(* Logix 5000 project; controller PLC_MCC1300_75F1 vendor 1 type 14 code 166 rev 32.11; software revision 32.04; part 76 of 83 *)
(* tags used below, declared in another part *)
   AUX_tCapsConveyor_NULL : UDT_CapsConveyor_ZC;
   CONST_tPlant : UDT_PLANT_CONSTANTS;
   M302SpeedUp_ALM : MAC_SpeedUp_ALM;
   M307ASpeedUp_ALM : MAC_SpeedUp_ALM;
   M30xTrimDeck : MAC_TrimmingDeck[5];
   M30xTrimWheel : MAC_TrimmingWheels[5];
   M312 : MAC_Conveyor_Single;
   TMP_dIndex : DINT;
   TMP_dIndexCapConv : DINT;
   TMP_dIndexConv : DINT;
   TMP_x : BOOL;
   TMP_xDummy : BOOL;
   xAlwaysOFF : BOOL;
   Z300_BufferPlate : UDT_LINE_BUFFER_PLATE;
   Z300_Conveyor : UDT_StandConv[29];
   Z300_Conveyor_HMW : MAC_Conveyor_ZC_HMW[29];
   Z300_LineTracking : UDT_LINE_TRACKING;
   Z301 : MAC_Zone_ML;
   Z301_ALM : MAC_Zone_ML_ALM;
   Z301_HMR : MAC_Zone_ML_HMR;
   Z301_HMW : MAC_Zone_ML_HMW;
(* MainProgram, continued *)

ROUTINE Tracking_Logic   (* structured text *)
   
   // Step advancement conveyor
   FOR TMP_dIndexConv:=0 TO CONST_tPlant.dNumOfConveyors - 1 DO
   	JSR(sbrTrackingConvStep,1,TMP_dIndexConv);
   	//reset conveyor tracking
   	FOR TMP_dIndexCapConv := 0 TO CONST_tPlant.dNumCapsConveyor - 1 DO
   		COP(AUX_tCapsConveyor_NULL,Z300_LineTracking.rgtTrkConv[TMP_dIndexConv].Cap[TMP_dIndexCapConv],1);
   	END_FOR;
   	Z300_LineTracking.rgtTrkConv[TMP_dIndexConv].dIndexCaps := 0;
   	Z300_LineTracking.rgtTrkConv[TMP_dIndexConv].xPlatePassageNext := 0;
   	Z300_LineTracking.rgtTrkConv[TMP_dIndexConv].xPlatePassagePrevious := 0;
   	Z300_LineTracking.rgtTrkConv[TMP_dIndexConv].xGlassPresence := 0;
   	Z300_LineTracking.rgtTrkConv[TMP_dIndexConv].xPlateConvPreviousNext := 0;
   	Z300_LineTracking.rgtTrkConv[TMP_dIndexConv].dTailPosition_cmm := 0;
   	Z300_LineTracking.rgtTrkConv[TMP_dIndexConv].dHeadPosition_cmm := 0;
   END_FOR;
   
   // Reset flag for tracking
   FOR TMP_dIndex:=0 TO CONST_tPlant.dMaxNumPlates - 1 DO
   	IF Z300_BufferPlate.rgtPlate[TMP_dIndex].tData.dLength_cmm <= 0 THEN
   		Z300_BufferPlate.rgtPlate[TMP_dIndex].tTracking.xHoldAdvancement := 0;
   		Z300_BufferPlate.rgtPlate[TMP_dIndex].tTracking.xNotConsConvTrk := 0;
   		Z300_BufferPlate.rgtPlate[TMP_dIndex].tTracking.xNotShownInScada := 0;
   	END_IF;
   END_FOR;
   
   // Tracking index not in convoy
   FOR TMP_dIndex:=0 TO CONST_tPlant.dMaxNumPlates - 1 DO
   	JSR(sbrTrackingIndexNotInConvoy,1,Z300_BufferPlate.rgtPlate[TMP_dIndex].tTracking);
   END_FOR;
   
   // Tracking shift
   JSR(sbrTrackingShift);
   
   // Plate presence convoy
   JSR(sbrTrackingConvPresence);
   
END_ROUTINE

ROUTINE Z301_Faults   (* ladder *)
   0: NOP();
   1: XIC(Z301.ST_xAlarmOff)MOV(0,Z301_ALM.rgxEmergency[0])MOV(0,Z301_ALM.rgxStoppingFault[0])MOV(0,Z301_ALM.rgxFault[0])MOV(0,Z301_ALM.rgxWarning[0])MOV(0,Z301_ALM.rgdFaultCode[0]);
   2: XIO(Z301.INPUT_x24VdcVoltageON)OTE(Z301_ALM.rgxStoppingFault[0].0);
   3: XIO(Z301.INPUT_xPowerSupply24VLogic1)OTE(Z301_ALM.rgxStoppingFault[0].3);
   4: XIO(Z301.INPUT_xPowerSupply24VLogic2)OTE(Z301_ALM.rgxStoppingFault[0].4);
   5: XIO(Z301.INPUT_xPowerSupply24VLogic3)OTE(Z301_ALM.rgxStoppingFault[0].5);
   6: XIO(Z301.INPUT_xPowerSupply24VDrive1)OTE(Z301_ALM.rgxStoppingFault[0].8);
   7: XIO(Z301.INPUT_xPowerSupply24VDrive2)OTE(Z301_ALM.rgxStoppingFault[0].9);
   8: XIO(Z301.INPUT_xEthernetSwitch24VON)OTE(Z301_ALM.rgxStoppingFault[0].13);
   9: XIO(Z301.INPUT_xPowerSupply400VDrive1)OTE(Z301_ALM.rgxStoppingFault[0].16);
   10: XIO(Z301.INPUT_xPowerSupply400VDrive2)OTE(Z301_ALM.rgxStoppingFault[0].17);
   11: XIO(Z301.INPUT_xPowerSupply230V_PLC1)OTE(Z301_ALM.rgxFault[0].0);
   12: XIO(Z301.INPUT_xPowerSupply230V_PLC2)OTE(Z301_ALM.rgxFault[0].1);
   13: XIC(Z301.INPUT_xEthernetSwitchFault)OTE(Z301_ALM.rgxFault[0].8);
   14: XIO(Z301.INPUT_xPowerSupply230V_Service)OTE(Z301_ALM.rgxWarning[0].0);
   15: XIO(Z301.INPUT_xMainEmergencyON)OTE(Z301_ALM.rgxEmergency[0].31);
   16: [XIC(Z301.INPUT_xEmergencyLocalization1) ,XIC(Z301_ALM.rgxEmergency[0].0) ]XIC(Z301_ALM.rgxEmergency[0].31)OTE(Z301_ALM.rgxEmergency[0].0);
   17: [XIC(Z301.INPUT_xEmergencyLocalization2) ,XIC(Z301_ALM.rgxEmergency[0].1) ]XIC(Z301_ALM.rgxEmergency[0].31)OTE(Z301_ALM.rgxEmergency[0].1);
   18: [XIC(Z301.INPUT_xEmergencyLocalization3) ,XIC(Z301_ALM.rgxEmergency[0].2) ]XIC(Z301_ALM.rgxEmergency[0].31)OTE(Z301_ALM.rgxEmergency[0].2);
   19: [XIC(Z301.INPUT_xEmergencyLocalization4) ,XIC(Z301_ALM.rgxEmergency[0].3) ]XIC(Z301_ALM.rgxEmergency[0].31)OTE(Z301_ALM.rgxEmergency[0].3);
   20: [XIC(Z301.INPUT_xEmergencyLocalization5) ,XIC(Z301_ALM.rgxEmergency[0].4) ]XIC(Z301_ALM.rgxEmergency[0].31)OTE(Z301_ALM.rgxEmergency[0].4);
   21: [XIC(Z301.INPUT_xEmergencyLocalization6) ,XIC(Z301_ALM.rgxEmergency[0].5) ]XIC(Z301_ALM.rgxEmergency[0].31)OTE(Z301_ALM.rgxEmergency[0].5);
   22: [XIC(Z301.INPUT_xEmergencyLocalization7) ,XIC(Z301_ALM.rgxEmergency[0].6) ]XIC(Z301_ALM.rgxEmergency[0].31)OTE(Z301_ALM.rgxEmergency[0].6);
   23: [XIC(Z301.INPUT_xEmergencyLocalization8) ,XIC(Z301_ALM.rgxEmergency[0].7) ]XIC(Z301_ALM.rgxEmergency[0].31)OTE(Z301_ALM.rgxEmergency[0].7);
END_ROUTINE

ROUTINE Z301_Logic   (* ladder *)
   // ##### MATCH #####
   0: NOP();
   // 24Vdc ON
   1: XIC(Z301.ST_xThisPlcActive)XIC(Z301.INPUT_x24VdcVoltageON)XIC(Z301.INPUT_xPowerSupply24VLogic1)XIC(Z301.INPUT_xPowerSupply24VLogic2)XIC(Z301.INPUT_xPowerSupply24VLogic3)XIC(Z301.INPUT_xEthernetSwitch24VON)XIC(Z301.INPUT_xPowerSupply24VDrive1)XIC(Z301.INPUT_xPowerSupply24VDrive2)TON(Z301.tmON_24Vdc,?,?);
   // 400Vac Drive ON
   2: XIC(Z301.ST_xThisPlcActive)XIC(Z301.INPUT_xPowerSupply400VDrive1)XIC(Z301.INPUT_xPowerSupply400VDrive2)TON(Z301.tmON_400Vca,?,?);
   3: XIC(Z301.ST_xThisPlcActive)XIC(Z301.INPUT_xMainEmergencyON)TON(Z301.tmON_EmergencyOK,?,?);
   // #####_ALARMS_#####
   4: NOP();
   5: XIC(Z301_HMW.xResetErrorRequest)[OTU(Z301_HMW.xResetErrorRequest) ,TOF(Z301.tmON_ResetAlarm,?,?) ];
   6: XIC(Z301.tmON_ResetAlarm.DN)OTE(Z301.ST_xAlarmOff);
   7: XIC(Z301.tmON_24Vdc.DN)XIC(Z301.tmON_400Vca.DN)XIC(Z301.tmON_EmergencyOK.DN)OTE(Z301.ST_xEnableControlError);
   8: JSR(Z301_Faults,0);
   // #####_HMI_LOGICS_#####
   9: NOP();
   // Thickness change mode enabled
   10: [XIC(Z301_HMW.xEnableChangeThick) [OTL(Z301_HMR.xChangeThickEnabled) ,OTU(Z301_HMW.xEnableChangeThick) ] ,XIC(Z301_HMW.xDisableChangeThick) [OTU(Z301_HMR.xChangeThickEnabled) ,OTU(Z301_HMW.xDisableChangeThick) ] ];
   // Enable/Disable automatic speed adjustment
   11: XIC(Z301_HMW.xEnDisableAutoSpeedAdjust)OTE(Z301_HMR.xAutoSpeedAdjustEnabled);
   // #####_STATUSES_#####
   12: NOP();
   13: [NEQ(Z301_ALM.rgxEmergency[0],0) ,NEQ(Z301_ALM.rgxStoppingFault[0],0) ,NEQ(Z301_ALM.rgxFault[0],0) ,NEQ(Z301_ALM.rgxWarning[0],0) ,NEQ(M302SpeedUp_ALM.rgxFault,0) ,NEQ(M302SpeedUp_ALM.rgxWarning,0) ,NEQ(M307ASpeedUp_ALM.rgxFault,0) ,NEQ(M307ASpeedUp_ALM.rgxWarning,0) ,XIC(M30xTrimDeck[0].ST_xMachineFault) ,XIC(M30xTrimDeck[1].ST_xMachineFault) ,XIC(M30xTrimDeck[2].ST_xMachineFault) ,XIC(M30xTrimDeck[3].ST_xMachineFault) ,XIC(M30xTrimDeck[4].ST_xMachineFault) ,XIC(M30xTrimWheel[0].ST_xMachineFaultOpSide) ,XIC(M30xTrimWheel[1].ST_xMachineFaultOpSide) ,XIC(M30xTrimWheel[2].ST_xMachineFaultOpSide) ,XIC(M30xTrimWheel[3].ST_xMachineFaultOpSide) ]OTE(Z301.ST_xZoneError);
   14: [XIC(Z300_Conveyor[0].ST_xStopMachineFault) ,XIC(Z300_Conveyor[1].ST_xStopMachineFault) ,XIC(Z300_Conveyor[2].ST_xStopMachineFault) ,XIC(Z300_Conveyor[3].ST_xStopMachineFault) ,XIC(Z300_Conveyor[4].ST_xStopMachineFault) ,XIC(Z300_Conveyor[5].ST_xStopMachineFault) ,XIC(Z300_Conveyor[6].ST_xStopMachineFault) ,XIC(Z300_Conveyor[7].ST_xStopMachineFault) ,XIC(Z300_Conveyor[8].ST_xStopMachineFault) ,XIC(Z300_Conveyor[9].ST_xStopMachineFault) ,XIC(Z300_Conveyor[10].ST_xStopMachineFault) ,XIC(Z300_Conveyor[11].ST_xStopMachineFault) ]XIC(Z301.ST_xCycleON)[TON(Z301.tmON_ConveyorsNotOK,?,?) ,XIC(Z301.tmON_ConveyorsNotOK.DN) OTE(Z301.ST_xConveyorsNotOK) ];
   // #####_ZONE_MODALITY_#####
   15: NOP();
   16: XIC(Z301_HMW.xManualModeReq)[OTL(Z301.ST_xSelManuMode) ,OTU(Z301.ST_xSelAutoMode) ,OTU(Z301_HMW.xManualModeReq) ];
   17: XIC(Z301_HMW.xAutoModeReq)[OTL(Z301.ST_xSelAutoMode) ,OTU(Z301.ST_xSelManuMode) ,OTU(Z301_HMW.xAutoModeReq) ];
   18: [XIC(Z301.ST_xConditionOKStopCycle) ,XIO(Z301.ST_xCycleON) ]OTE(Z301.ST_xManualModeConditionOK);
   19: XIC(Z301.ST_xSelManuMode)[XIO(Z301.ST_xManuModeAccepted) OTE(Z301.ST_xManuModeReq) ,[XIC(Z301.ST_xManualModeConditionOK) ,XIC(Z301.ST_xManuModeAccepted) ] [OTE(Z301.ST_xManuModeAccepted) ,ONS(Z301.OSR_xManualAccepted) OTE(Z301.OS_xManualAccepted) ] ];
   20: XIO(Z301.ST_xManuModeAccepted)[XIC(Z301.ST_xSelAutoMode) ,XIC(Z301.ST_xAutoModeAccepted) ][OTE(Z301.ST_xAutoModeAccepted) ,ONS(Z301.OSR_xAutoAccepted) OTE(Z301.OS_xAutoAccepted) ];
   21: XIC(Z301.OS_xManualAccepted)[OTL(Z300_Conveyor_HMW[0].xEnableDisableManualCommand) ,OTL(Z300_Conveyor_HMW[5].xEnableDisableManualCommand) ,OTL(Z300_Conveyor_HMW[6].xEnableDisableManualCommand) ,OTL(Z300_Conveyor_HMW[7].xEnableDisableManualCommand) ,OTL(Z300_Conveyor_HMW[8].xEnableDisableManualCommand) ,OTL(Z300_Conveyor_HMW[11].xEnableDisableManualCommand) ];
   22: XIC(Z301.OS_xAutoAccepted)[OTU(Z300_Conveyor_HMW[0].xEnableDisableManualCommand) ,OTU(Z300_Conveyor_HMW[5].xEnableDisableManualCommand) ,OTU(Z300_Conveyor_HMW[6].xEnableDisableManualCommand) ,OTU(Z300_Conveyor_HMW[7].xEnableDisableManualCommand) ,OTU(Z300_Conveyor_HMW[8].xEnableDisableManualCommand) ,OTU(Z300_Conveyor_HMW[11].xEnableDisableManualCommand) ];
   // M301 Manual Command Enabled
   23: XIC(Z300_Conveyor_HMW[0].xEnableDisableManualCommand)[OTE(Z300_Conveyor_HMW[1].xEnableDisableManualCommand) ,OTE(Z300_Conveyor_HMW[2].xEnableDisableManualCommand) ,OTE(Z300_Conveyor_HMW[3].xEnableDisableManualCommand) ,OTE(Z300_Conveyor_HMW[4].xEnableDisableManualCommand) ];
   // M312 Manual Command Enabled
   24: XIC(Z300_Conveyor_HMW[8].xEnableDisableManualCommand)[OTE(Z300_Conveyor_HMW[9].xEnableDisableManualCommand) ,OTE(Z300_Conveyor_HMW[10].xEnableDisableManualCommand) ];
   // M301 Manual Command Enabled
   25: XIC(Z300_Conveyor_HMW[0].rgxMan.xAllFwd)[OTE(Z300_Conveyor_HMW[1].rgxMan.xAllFwd) ,OTE(Z300_Conveyor_HMW[2].rgxMan.xAllFwd) ,OTE(Z300_Conveyor_HMW[3].rgxMan.xAllFwd) ,OTE(Z300_Conveyor_HMW[4].rgxMan.xAllFwd) ];
   // M312 Manual Command Enabled
   26: XIC(Z300_Conveyor_HMW[8].rgxMan.xAllFwd)[OTE(Z300_Conveyor_HMW[9].rgxMan.xAllFwd) ,OTE(Z300_Conveyor_HMW[10].rgxMan.xAllFwd) ];
   // M301 Manual Command Enabled
   27: XIC(Z300_Conveyor_HMW[0].rgxMan.xAllBwd)[OTE(Z300_Conveyor_HMW[1].rgxMan.xAllBwd) ,OTE(Z300_Conveyor_HMW[2].rgxMan.xAllBwd) ,OTE(Z300_Conveyor_HMW[3].rgxMan.xAllBwd) ,OTE(Z300_Conveyor_HMW[4].rgxMan.xAllBwd) ];
   // M312 Manual Command Enabled
   28: XIC(Z300_Conveyor_HMW[8].rgxMan.xAllBwd)[OTE(Z300_Conveyor_HMW[9].rgxMan.xAllBwd) ,OTE(Z300_Conveyor_HMW[10].rgxMan.xAllBwd) ];
   // #####_START/STOP ZONE_#####
   29: NOP();
   30: XIC(Z301_HMW.xStartCycleRequest)[OTE(Z301.OS_xStartCycle) ,OTU(Z301_HMW.xStartCycleRequest) ];
   31: XIC(Z301_HMW.xStopCycleRequest)[OTE(Z301.OS_xStopCycle) ,OTU(Z301_HMW.xStopCycleRequest) ];
   32: XIC(xAlwaysOFF)TON(Z301.tmON_ForceStop,?,?);
   33: [XIC(Z301_HMW.xForceStopCycle) ,XIC(Z301.tmON_ForceStop.DN) ONS(Z301.OSR_xForceStopCycle) ][OTE(Z301.OS_xForceStopCycle) ,OTU(Z301_HMW.xForceStopCycle) ];
   34: XIC(Z301.ST_xCycleON)XIC(Z301.ST_xConveyorsNotOK)OTE(Z301.ST_xStopCycleReqForFaults);
   35: XIC(Z301.ST_xCycleON)XIC(Z301.ST_xStopCycleReqForFaults)[TON(Z301.tmON_StopCycleForFaults,?,?) ,XIC(Z301.tmON_StopCycleForFaults.DN) OTE(Z301.ST_xStopCycleAcceptForFaults) ];
   36: XIO(Z300_Conveyor[0].ST_xManualCmdEnabled)XIO(Z300_Conveyor[1].ST_xManualCmdEnabled)XIO(Z300_Conveyor[2].ST_xManualCmdEnabled)XIO(Z300_Conveyor[3].ST_xManualCmdEnabled)XIO(Z300_Conveyor[4].ST_xManualCmdEnabled)XIO(Z300_Conveyor[5].ST_xManualCmdEnabled)XIO(Z300_Conveyor[6].ST_xManualCmdEnabled)XIO(Z300_Conveyor[7].ST_xManualCmdEnabled)XIO(Z300_Conveyor[8].ST_xManualCmdEnabled)XIO(Z300_Conveyor[9].ST_xManualCmdEnabled)XIO(Z300_Conveyor[10].ST_xManualCmdEnabled)XIO(Z300_Conveyor[11].ST_xManualCmdEnabled)XIO(Z300_Conveyor[0].ST_xFaulted)XIO(Z300_Conveyor[1].ST_xFaulted)XIO(Z300_Conveyor[2].ST_xFaulted)XIO(Z300_Conveyor[3].ST_xFaulted)XIO(Z300_Conveyor[4].ST_xFaulted)XIO(Z300_Conveyor[5].ST_xFaulted)XIO(Z300_Conveyor[6].ST_xFaulted)XIO(Z300_Conveyor[7].ST_xFaulted)XIO(Z300_Conveyor[8].ST_xFaulted)XIO(Z300_Conveyor[9].ST_xFaulted)XIO(Z300_Conveyor[10].ST_xFaulted)XIO(Z300_Conveyor[11].ST_xFaulted)OTE(TMP_x);
   37: XIC(Z301.ST_xAutoModeAccepted)XIO(Z301.ST_xStopCycleAcceptForFaults)XIO(Z301.ST_xStopCycleForSaturation)XIC(Z301.tmON_24Vdc.DN)XIC(Z301.tmON_400Vca.DN)XIC(Z301.tmON_EmergencyOK.DN)XIC(TMP_x)OTE(Z301.ST_xConditionOkCycleON);
   38: [XIC(Z301.OS_xStartCycle) ,XIC(Z301.ST_xStartCycleRequest) ]XIC(Z301.ST_xConditionOkCycleON)[XIO(Z301.ST_xCycleON) ,XIC(Z301.ST_xStopCycleRequest) ]XIO(Z301.OS_xStopCycle)OTE(Z301.ST_xStartCycleRequest);
   39: [XIC(Z301.OS_xStopCycle) ,XIC(Z301.ST_xManuModeReq) ,XIC(Z301.ST_xStopCycleRequest) ]XIC(Z301.ST_xCycleON)XIO(Z301.ST_xStartCycleRequest)OTE(Z301.ST_xStopCycleRequest);
   40: XIC(Z300_Conveyor[0].ST_xStopCycleConditionOK)XIC(Z300_Conveyor[1].ST_xStopCycleConditionOK)XIC(Z300_Conveyor[2].ST_xStopCycleConditionOK)XIC(Z300_Conveyor[3].ST_xStopCycleConditionOK)XIC(Z300_Conveyor[4].ST_xStopCycleConditionOK)XIC(Z300_Conveyor[5].ST_xStopCycleConditionOK)XIC(Z300_Conveyor[6].ST_xStopCycleConditionOK)XIC(Z300_Conveyor[7].ST_xStopCycleConditionOK)XIC(Z300_Conveyor[8].ST_xStopCycleConditionOK)XIC(Z300_Conveyor[9].ST_xStopCycleConditionOK)XIC(Z300_Conveyor[10].ST_xStopCycleConditionOK)XIC(Z300_Conveyor[11].ST_xStopCycleConditionOK)XIC(Z300_Conveyor[12].ST_xStopCycleConditionOK)XIC(Z300_Conveyor[13].ST_xStopCycleConditionOK)XIC(Z300_Conveyor[14].ST_xStopCycleConditionOK)XIC(Z300_Conveyor[15].ST_xStopCycleConditionOK)XIC(Z300_Conveyor[16].ST_xStopCycleConditionOK)XIC(Z300_Conveyor[17].ST_xStopCycleConditionOK)XIC(Z300_Conveyor[18].ST_xStopCycleConditionOK)XIC(M30xTrimDeck[0].ST_xConditionOKStopCycle)XIC(M30xTrimDeck[1].ST_xConditionOKStopCycle)XIC(M30xTrimDeck[2].ST_xConditionOKStopCycle)XIC(M30xTrimDeck[3].ST_xConditionOKStopCycle)XIC(M30xTrimDeck[4].ST_xConditionOKStopCycle)XIC(M30xTrimWheel[0].ST_xConditionOKStopCycle)XIC(M30xTrimWheel[1].ST_xConditionOKStopCycle)XIC(M30xTrimWheel[2].ST_xConditionOKStopCycle)XIC(M30xTrimWheel[3].ST_xConditionOKStopCycle)XIC(M30xTrimWheel[4].ST_xConditionOKStopCycle)OTE(Z301.ST_xConditionOKStopCycle);
   41: XIC(Z301.ST_xStopCycleRequest)XIC(Z301.ST_xConditionOKStopCycle)OTE(Z301.ST_xStopCycleAccepted);
   42: [XIC(Z301.ST_xStartCycleRequest) ,XIC(Z301.ST_xCycleON) ]XIC(Z301.ST_xConditionOkCycleON)XIO(Z301.OS_xForceStopCycle)XIO(Z301.ST_xStopCycleAccepted)[TON(Z301.tmON_Cycle,?,?) ,XIC(Z301.tmON_Cycle.DN) OTE(Z301.ST_xCycleON) ];
   43: XIC(Z301.ST_xCycleON)XIO(Z301.ST_xManuModeReq)XIO(Z301.ST_xStopCycleRequest)XIO(Z301.ST_xStopCycleReqForFaults)OTE(Z301.ST_xConditionOkPhaseAdvancement);
   // #####_CLEANING_#####
   44: NOP();
   45: [XIC(Z301_HMW.xStartCleanZoneRequest) ,XIC(Z301.ST_xReqCleaningWrongLength) ,XIC(Z301.ST_xReqCleaningMissSnap) ,XIC(Z301.ST_xReqCleaningBufferOverflow) ][OTL(Z301.ST_xReqCleaning) ,OTU(Z301_HMW.xStartCleanZoneRequest) ];
   46: XIC(Z301_HMW.xStopCleanZoneRequest)[OTE(TMP_xDummy) ,OTU(Z301_HMW.xStopCleanZoneRequest) ];
   47: [XIC(Z301.ST_xCleaningAccepted) ,XIC(TMP_xDummy) ]OTU(Z301.ST_xReqCleaning);
   48: XIC(Z301.ST_xCleaningAccepted)[[XIC(TMP_xDummy) ,XIC(Z301.ST_xReqCleaningMissSnap) ,XIC(Z301.ST_xReqCleaningBufferOverflow) ] OTU(Z301.ST_xCleaningAccepted) ,OTU(Z301.ST_xReqCleaningCPUSwitching) ,OTU(Z301.ST_xReqCleaningWrongLength) ,OTU(Z301.ST_xReqCleaningMissSnap) ,OTU(Z301.ST_xReqCleaningBufferOverflow) ];
   49: XIC(Z300_Conveyor[0].tIN_Zone.xCleanZoneAccepted)[OTE(Z300_Conveyor_HMW[0].xLocalCleaningRequest) ,MOV(0,Z301.AUX_dStartIndexCleaning) ];
   // M301 Cleaning Enabled
   50: XIC(Z300_Conveyor_HMW[0].xLocalCleaningRequest)XIC(Z300_Conveyor[0].tIN_Zone.xCleanZoneAccepted)[OTE(Z300_Conveyor_HMW[1].xLocalCleaningRequest) ,OTE(Z300_Conveyor_HMW[2].xLocalCleaningRequest) ,OTE(Z300_Conveyor_HMW[3].xLocalCleaningRequest) ,OTE(Z300_Conveyor_HMW[4].xLocalCleaningRequest) ];
   51: XIC(Z300_Conveyor_HMW[4].xLocalCleaningRequest)XIC(Z300_Conveyor[0].tIN_Zone.xCleanZoneAccepted)OTE(Z300_Conveyor_HMW[5].xLocalCleaningRequest);
   52: XIC(Z300_Conveyor_HMW[5].xLocalCleaningRequest)XIC(Z300_Conveyor[0].tIN_Zone.xCleanZoneAccepted)OTE(Z300_Conveyor_HMW[6].xLocalCleaningRequest);
   53: XIC(Z300_Conveyor_HMW[6].xLocalCleaningRequest)XIC(Z300_Conveyor[0].tIN_Zone.xCleanZoneAccepted)OTE(Z300_Conveyor_HMW[7].xLocalCleaningRequest);
